     (* Datenbaustein Testen *)
     #rTEST_DB := TEST_DB(DB_NUMBER := #_pt.DBNr // IN: WORD
                        ,DB_LENGTH => #DB_LENGTH // OUT: WORD
                        ,WRITE_PROT => #WRITE_PROT // OUT: BOOL
                        ); // INT
     (* Ende wenn Test-DB <> 0 = Fehler *)
     IF #rTEST_DB <> 0 THEN RETURN; END_IF;
     (* Ende wenn DB zu klein *) 
     IF WORD_TO_INT(#DB_LENGTH)/4 < #size THEN RETURN; END_IF;

     #Adr := DWORD_TO_INT(SHR(IN:=SHL(IN:=#_pt.Adr,N:=8),N:=11));

     (* at first we calualte the arithmetic average of the array *)

     #stop := (#size - 1) / 1;     // (size -SIZEOF(pt)) / SIZEOF(pt);
     #avg := DWORD_TO_REAL(WORD_TO_BLOCK_DB(#_pt.DBNr).DD(#Adr+0));
     FOR #i := 1 TO #stop DO
         #avg := #avg + DWORD_TO_REAL(WORD_TO_BLOCK_DB(#_pt.DBNr).DD(#Adr+#i*4));
     END_FOR;
     #avg := #avg / (#stop + 1);

     (* in a second run we calculate the variance of the array *)

     #_var := (DWORD_TO_REAL(WORD_TO_BLOCK_DB(#_pt.DBNr).DD(#Adr+0)) - #avg) ** 2;
     FOR #i := 1 TO #stop DO
         #_var := #_var + ((DWORD_TO_REAL(WORD_TO_BLOCK_DB(#_pt.DBNr).DD(#Adr+#i*4)) - #avg) ** 2);
     END_FOR;
     #_var := #_var / #stop;

     (* standard deviation is simply the square root of the variance *)

     #sdv := SQRT(#_var);

   (*
   (* standard deviation is simply the square root of the variance *)

   array_sdv := SQRT(array_var(pt, size));
   *)

   (* revision history
   hm  1.4.2007        rev 1.0
       function created

   hm  16. mar. 2008   rev 1.1
       changed type of input size to uint

   *)
END_FUNCTION_BLOCK

FUNCTION_BLOCK "ARRAY_SPR"   // FB18, SCL
TITLE = ARRAY_SPR
{ S7_Optimized_Access := 'FALSE' }
AUTHOR : hugo
FAMILY : ARFUNCT
NAME : AR_SPR
VERSION : 1.1
// this function will calculate the spread of a given array.
// the function needs to be called:    array_spr(adr("array"),sizeof("array"));
// for example: spread of [12,0,4,1,7] is 12 - 0 = 12.
// because this function works with pointers its very time efficient and it needs no extra memory.
   VAR_INPUT
      pt : Pointer;
      _pt AT pt : Struct
         DBNr : Word;
         Adr : DWord;
      END_STRUCT;
      size : Int;
   END_VAR
   VAR_OUTPUT
      spr : Real;
   END_VAR
   VAR_TEMP
      i : Int;
      stop : Int;
      array_max : Real;
      array_min : Real;
      Adr : Int;
      DB_LENGTH : Word;
      WRITE_PROT : Bool;
      rTEST_DB : Int;
   END_VAR
BEGIN


     (* Datenbaustein Testen *)
     #rTEST_DB := TEST_DB(DB_NUMBER := #_pt.DBNr // IN: WORD
                        ,DB_LENGTH => #DB_LENGTH // OUT: WORD
                        ,WRITE_PROT => #WRITE_PROT // OUT: BOOL
                        ); // INT
     (* Ende wenn Test-DB <> 0 = Fehler *)
     IF #rTEST_DB <> 0 THEN RETURN; END_IF;
     (* Ende wenn DB zu klein *) 
     IF WORD_TO_INT(#DB_LENGTH)/4 < #size THEN RETURN; END_IF;

     #Adr := DWORD_TO_INT(SHR(IN:=SHL(IN:=#_pt.Adr,N:=8),N:=11));

     (* Berechnung *)
     #stop := (#size - #size / #size);
     #array_min := DWORD_TO_REAL(WORD_TO_BLOCK_DB(#_pt.DBNr).DD(#Adr+0));
     #array_max := DWORD_TO_REAL(WORD_TO_BLOCK_DB(#_pt.DBNr).DD(#Adr+0));
     FOR #i := 1 TO #stop DO
         IF DWORD_TO_REAL(WORD_TO_BLOCK_DB(#_pt.DBNr).DD(#Adr+#i*4)) > #array_max THEN 
             #array_max := DWORD_TO_REAL(WORD_TO_BLOCK_DB(#_pt.DBNr).DD(#Adr+#i*4));
         ELSIF DWORD_TO_REAL(WORD_TO_BLOCK_DB(#_pt.DBNr).DD(#Adr+#i*4)) < #array_min THEN 
             #array_min := DWORD_TO_REAL(WORD_TO_BLOCK_DB(#_pt.DBNr).DD(#Adr+#i*4));
         END_IF;
     END_FOR;
     #spr := #array_max - #array_min;

   (* revision history
   hm  2. oct. 2006    rev 1.0
       original version

   hm  16. mar. 2008   rev 1.1
       changed type of input size to uint

   *)
END_FUNCTION_BLOCK

FUNCTION_BLOCK "ARRAY_SUM"   // FB19, SCL
TITLE = ARRAY_SUM
{ S7_Optimized_Access := 'FALSE' }
AUTHOR : hugo
FAMILY : ARFUNCT
NAME : AR_SUM
VERSION : 1.1
// this function will calculate the sum of a given array.
   VAR_INPUT
      pt : Pointer;
      _pt AT pt : Struct
         DBNr : Word;
         Adr : DWord;
      END_STRUCT;
      size : Int;
   END_VAR
   VAR_OUTPUT
      sum : Real;
   END_VAR
   VAR_TEMP
      i : Int;
      Adr : Int;
      DB_LENGTH : Word;
      WRITE_PROT : Bool;
      rTEST_DB : Int;
   END_VAR
BEGIN


     (* Datenbaustein Testen *)
     #rTEST_DB := TEST_DB(DB_NUMBER := #_pt.DBNr // IN: WORD
                        ,DB_LENGTH => #DB_LENGTH // OUT: WORD
                        ,WRITE_PROT => #WRITE_PROT // OUT: BOOL
                        ); // INT
     (* Ende wenn Test-DB <> 0 = Fehler *)
     IF #rTEST_DB <> 0 THEN RETURN; END_IF;
     (* Ende wenn DB zu klein *) 
     IF WORD_TO_INT(#DB_LENGTH)/4 < #size THEN RETURN; END_IF;

     #Adr := DWORD_TO_INT(SHR(IN:=SHL(IN:=#_pt.Adr,N:=8),N:=11));

     (* Berechnung *)
     #sum := DWORD_TO_REAL(WORD_TO_BLOCK_DB(#_pt.DBNr).DD(#Adr+0));
     FOR #i := 1 TO #size-1 DO
         #sum := #sum + DWORD_TO_REAL(WORD_TO_BLOCK_DB(#_pt.DBNr).DD(#Adr+#i*4));
     END_FOR;

   (* revision history
   hm  2. oct. 2006    rev 1.0
       function created

   hm  16. mar. 2008   rev 1.1
       changed type of input size to uint

   *)
END_FUNCTION_BLOCK

FUNCTION_BLOCK "ARRAY_TREND"   // FB20, SCL
TITLE = ARRAY_TREND
{ S7_Optimized_Access := 'FALSE' }
AUTHOR : hugo
FAMILY : ARFUNCT
NAME : AR_TREND
VERSION : 1.3
// this function will calculate the trend of a given array.
// trend will calculate the avg of the first half of the array and then the avg of the second half, trend = avg2 - avg1.
// for example:  [0,1,4,5,3,4,6,3] = 4 - 2.5 = 1.5
// the function needs to be called:    array_trend(adr("array"),sizeof("array"));
// because this function works with pointers its very time efficient and it needs no extra memory.
// 
// uses: EVEN [FC76]
   VAR_INPUT
      pt : Pointer;
      _pt AT pt : Struct
         DBNr : Word;
         Adr : DWord;
      END_STRUCT;
      size : Int;
   END_VAR
   VAR_OUTPUT
      trend : Real;
   END_VAR
   VAR_TEMP
      i : Int;
      stop : Int;
      stop2 : Int;
      x : Real;
      Adr : Int;
      DB_LENGTH : Word;
      WRITE_PROT : Bool;
      rTEST_DB : Int;
   END_VAR
BEGIN


   (* Datenbaustein Testen *)
   #rTEST_DB := TEST_DB(DB_NUMBER := #_pt.DBNr, DB_LENGTH => #DB_LENGTH, WRITE_PROT => #WRITE_PROT);
   (* Ende wenn Test-DB <> 0 = Fehler *)
   IF #rTEST_DB <> 0 THEN RETURN; END_IF;
   (* Ende wenn DB zu klein *) 
   IF WORD_TO_INT(#DB_LENGTH)/4 < #size THEN RETURN; END_IF;

   #Adr := DWORD_TO_INT(SHR(IN:=SHL(IN:=#_pt.Adr,N:=8),N:=11));

   #stop := #size - 1;
   #stop2 := #stop / 2;
   FOR #i := 0 TO #stop2 DO #x := #x - DWORD_TO_REAL(WORD_TO_BLOCK_DB(#_pt.DBNr).DD(#Adr+#i*4)); END_FOR;
   IF "EVEN"(#stop) THEN
       FOR #i := #stop2 TO #stop DO #x := #x + DWORD_TO_REAL(WORD_TO_BLOCK_DB(#_pt.DBNr).DD(#Adr+#i*4)); END_FOR;
   ELSE
       FOR #i := #stop2 + 1 TO #stop DO #x := #x + DWORD_TO_REAL(WORD_TO_BLOCK_DB(#_pt.DBNr).DD(#Adr+#i*4)); END_FOR;
   END_IF;
   #trend := #x / INT_TO_REAL(#stop2 + 1);


   (* revision history
   hm  2 oct 2007  rev 1.0
       original version

   hm  12 dec 2007 rev 1.1
       changed code for better performance

   hm  16. mar. 2008   rev 1.2
       changed type of input size to uint

   hm  10. mar. 2009   rev 1.3
       added type conversions for compatibility reasons
   *)
END_FUNCTION_BLOCK

FUNCTION_BLOCK "ARRAY_VAR"   // FB21, SCL
TITLE = ARRAY_VAR
{ S7_Optimized_Access := 'FALSE' }
AUTHOR : hugo
FAMILY : ARFUNCT
NAME : AR_VAR
VERSION : 1.3
// this function will calculate the variance of a given array.
// the function needs to be called:    array_var(adr("array"),sizeof("array"));
// because this function works with pointers its very time efficient and it needs no extra memory.
   VAR_INPUT
      pt : Pointer;
      _pt AT pt : Struct
         DBNr : Word;
         Adr : DWord;
      END_STRUCT;
      size : Int;
   END_VAR
   VAR_OUTPUT
      _var : Real;
   END_VAR
   VAR_TEMP
      i : Int;
      stop : Int;
      avg : Real;
      Adr : Int;
      DB_LENGTH : Word;
      WRITE_PROT : Bool;
      rTEST_DB : Int;
   END_VAR
BEGIN


   (* Datenbaustein Testen *)
   #rTEST_DB := TEST_DB(DB_NUMBER := #_pt.DBNr, DB_LENGTH => #DB_LENGTH, WRITE_PROT => #WRITE_PROT);
   (* Ende wenn Test-DB <> 0 = Fehler *)
   IF #rTEST_DB <> 0 THEN RETURN; END_IF;
   (* Ende wenn DB zu klein *) 
   IF WORD_TO_INT(#DB_LENGTH)/4 < #size THEN RETURN; END_IF;

   #Adr := DWORD_TO_INT(SHR(IN:=SHL(IN:=#_pt.Adr,N:=8),N:=11));

   (* at first we calualte the arithmetic average of the array *)

   #stop := #size - 1;
   #avg := DWORD_TO_REAL(WORD_TO_BLOCK_DB(#_pt.DBNr).DD(#Adr+0));
   FOR #i := 1 TO #stop DO
       #avg := #avg + DWORD_TO_REAL(WORD_TO_BLOCK_DB(#_pt.DBNr).DD(#Adr+#i*4));
   END_FOR;
   #avg := #avg / (#stop + 1);

   (* in a second run we calculate the variance of the array *)

   #_var := (DWORD_TO_REAL(WORD_TO_BLOCK_DB(#_pt.DBNr).DD(#Adr+0)) - #avg) * (DWORD_TO_REAL(WORD_TO_BLOCK_DB(#_pt.DBNr).DD(#Adr+0)) - #avg);
   FOR #i := 1 TO #stop DO
       #_var := #_var + (DWORD_TO_REAL(WORD_TO_BLOCK_DB(#_pt.DBNr).DD(#Adr+#i*4)) - #avg) * (DWORD_TO_REAL(WORD_TO_BLOCK_DB(#_pt.DBNr).DD(#Adr+#i*4)) - #avg);
   END_FOR;
   #_var := #_var / INT_TO_REAL(#stop);


   (* revision history
   hm  1.4.2007    rev 1.0
       function created

   hm  12.12.2007  rev 1.1
       changed code for better performance

   hm  16. mar. 2008   rev 1.2
       changed type of input size to uint

   hm  10. mar. 2009   rev 1.3
       added type conversions for compatibility reasons
   *)
END_FUNCTION_BLOCK

FUNCTION_BLOCK "IS_SORTED"   // FB22, SCL
TITLE = IS_SORTED
{ S7_Optimized_Access := 'FALSE' }
AUTHOR : hugo
FAMILY : ARFUNCT
NAME : ARSORTED
VERSION : 1.1
// this function will return true if the given array is sorted in an ascending order.
// the function needs to be called:    array_sorted(adr("array"),sizeof("array"));
// because this function works with pointers its very time efficient and it needs no extra memory.
   VAR_INPUT
      pt : Pointer;
      _pt AT pt : Struct
         DBNr : Word;
         Adr : DWord;
      END_STRUCT;
      size : Int;
   END_VAR
   VAR_OUTPUT
      SORTED : Bool;
   END_VAR
   VAR
      stop : Int;
      i : Int;
      Adr : Int;
      DB_LENGTH : Word;
      WRITE_PROT : Bool;
      rTEST_DB : Int;
   END_VAR
BEGIN


   #SORTED := FALSE;

   (* Datenbaustein Testen *)
   #rTEST_DB := TEST_DB(DB_NUMBER := #_pt.DBNr // IN: WORD
                      ,DB_LENGTH => #DB_LENGTH // OUT: WORD
                      ,WRITE_PROT => #WRITE_PROT // OUT: BOOL
                      ); // INT
   (* Ende wenn Test-DB <> 0 = Fehler *)
   IF #rTEST_DB <> 0 THEN RETURN; END_IF;
   (* Ende wenn DB zu klein *) 
   IF WORD_TO_INT(#DB_LENGTH)/4 < #size THEN RETURN; END_IF;

   #Adr := DWORD_TO_INT(SHR(IN:=SHL(IN:=#_pt.Adr,N:=8),N:=11));

   #stop := #size - 2;   //WORD_TO_INT(SHR(IN:=INT_TO_WORD(size),N:=2))-2;
   FOR #i := 0 TO #stop DO
       IF DWORD_TO_REAL(WORD_TO_BLOCK_DB(#_pt.DBNr).DD(#Adr+#i*4)) > DWORD_TO_REAL(WORD_TO_BLOCK_DB(#_pt.DBNr).DD(#Adr+(#i+1)*4)) THEN
           #SORTED := FALSE;
           RETURN;
       END_IF;
   END_FOR;
   #SORTED := TRUE;

   (* revision history

   hm  29. mar. 2008   rev 1.0
       original version

   hm  4. apr. 2008    rev 1.1
       added type conversion to avoid warnings under codesys 3.0
   *)
END_FUNCTION_BLOCK

FUNCTION_BLOCK "STIME"   // FB64, SCL
TITLE = STIME
{ S7_Optimized_Access := 'FALSE' }
AUTHOR : dalbi
FAMILY : MEASURE
NAME : STIME
VERSION : 1.4
// this function block makes sure that the timer of a siemens sps counts from 0 - 2^32-1.
   VAR_OUTPUT
      tx : DWord;
      at_tx AT tx : Array[0..31] of Bool;
   END_VAR
   VAR
      last_time : DWord;
      bit31 : Bool;
      init : Bool := TRUE;
   END_VAR
   VAR_TEMP
      TOP_SI : Struct
         EV_CLASS : Byte;
         EV_NUM : Byte;
         PRIORITY : Byte;
         NUM : Byte;
         TYP2_3 : Byte;
         TYP1 : Byte;
         ZI1 : Word;
         ZI2_3 : DWord;
      END_STRUCT;
      START_UP_SI : Struct
         EV_CLASS : Byte;
         EV_NUM : Byte;
         PRIORITY : Byte;
         NUM : Byte;
         TYP2_3 : Byte;
         TYP1 : Byte;
         ZI1 : Word;
         ZI2_3 : DWord;
      END_STRUCT;
      ERR : Int;
   END_VAR
BEGIN


   (* this FB is only necessary for siemens sps
   the siemens sps timer counts from 0 to 2^31-1 and starts at 0 sfter overrun.
   this means that the bit 31 (the highest bit ) will never be used and therefore
   a problem arises when t2 - t1 is checked.
   t2 - t1 is always valid also in an timer overrun situation where the time t1 is very high and t2 is very low.
   the result of the subtraction t2 - t1 however is still valid.
   this calculation does not work for soiemens because the highest bit is not used.

   this module stores the highest bit, changes the highest bit at every overrun occurence and stuffs ther highest bit in the output.
   the output is then used by t_plc_us and t_plc_ms.

   the correction needs and fb and not a function because the value of the highest bit has to be stored.

   do never use this function block in a codesys environment. the timer in codesys is correct and runs from 0 to 2^32-1
   *)

   (* read actual startup info *)
   (* OB1_SCAN_1  BYTE  -  B#16#01: Abschluss des Neustarts (Warmstarts)
                        -  B#16#02: Abschluss des Wiederanlaufs
                        -  B#16#03: Abschluss des freien Zyklus
                        -  B#16#04: Abschluss des Kaltstarts
                        -  B#16#05: Erster OB 1-Zyklus der neuen Master-CPU nach 
                                    Master-Reserve-Umschaltung und STOP des 
                                    bisherigen Masters *)

   #ERR := RD_SINFO (TOP_SI => #TOP_SI, START_UP_SI => #START_UP_SI);

   (* reset last_time on system startup *)
   IF #TOP_SI.EV_NUM = 1 OR #TOP_SI.EV_NUM = 2 OR #TOP_SI.EV_NUM = 4 OR NOT #init THEN 
       #last_time := 0;
       #bit31 := false;
       #init := true;
   END_IF;

   (* read the system timer *)
   #tx := DINT_TO_DWORD(T_CONV(TIME_TCK()));

   (* check for overrun *)
   IF DWORD_TO_DINT(#tx) < DWORD_TO_DINT(#last_time) THEN
       (* an overrun has occured, change the value of the highest bit *)
       #bit31 := NOT #bit31;
   END_IF;

   (* stuff the highest bit into the timer value *)
   #at_tx[7] := #bit31;

   (* remember the last system time for the next overrun check *)
   #last_time := #tx;


   (* revision history
   DA  14.9.2007 rev 1.0
     original version

   DA  24.2.2008 rev 1.1
     added self reset on system startup

   DA   2.5.2008 rev 1.2
     corect a problem running under OB35

   DA  12.3.2009 rev 1.3
     corect a problem run on different CPUs

   DA  22.12.2009 rev 1.4
     corect a problem on startup
   *)
END_FUNCTION_BLOCK

FUNCTION "T_PLC_MS" : DWord   // FC64, SCL
TITLE = T_PLC_MS
{ S7_Optimized_Access := 'FALSE' }
AUTHOR : hugo
FAMILY : MEASURE
NAME : T_PLC_MS
VERSION : 1.2
// T_PLC_MS reads the internal PLC timer and return the time, it has the advantage to be able to set a debug mode 
// and speed up the counter to test the plc timer overrun which occurs every 50 days respectively 25 days at siemens S7
// this routine also allows to correct the behavior of s7 where the internal plc counter will not count all 32 bits.
// 
// uses: STIME [FB64],IDB_STIME [DB64]
BEGIN


   "IDB_STIME"(); 
   #T_PLC_MS := "IDB_STIME".tx; 
   (* hier muss die korrektur für step7 stattfinden
   plctime muss den vollen wertebereich von time ausnutzen:
   wenn bei step7 time -24tage bis plus 24 tage ist dann muss der timer auch beim überlauf auf -24tage springen 
   und auf keinen fall auf 0 !!!!
   für siemens muss ein weiterer fb im main eingebunden werden der sicherstellt das alle 32 bits durchgezählt werden.
   es kann nur ein fb sein den er muss sich das oberste (32te) bit merken.
   oder etwa spring s7 bei überlauf auf -24 tage????? dann wäre keine korrektur nötig.
   *)
   IF "debug" THEN
       #T_PLC_MS := DINT_TO_DWORD((DWORD_TO_DINT(SHL(IN:=#T_PLC_MS,N:="N") OR SHL(IN:=DWORD#1,N:="N"))-1) + DWORD_TO_DINT("offset_1"));
   END_IF;


   (* revision history
   hm  14.9.2007   rev 1.0
       original version

   hm  12. nov 2007    rev 1.1
       added temporaray variable tx because some compilers could not handle time() as an argument

   hm  16. nov. 2008   rev 1.2
       initialized constants with 0 for compatibility reasons
   *)
END_FUNCTION

FUNCTION "EVEN" : Bool   // FC76, SCL
TITLE = EVEN
{ S7_Optimized_Access := 'FALSE' }
AUTHOR : hugo
FAMILY : MATH
NAME : EVEN
VERSION : 1.2
// this function chacks an input for even value
// the output is true if the input is even.
   VAR_INPUT
      in : DInt;
   END_VAR
   VAR_TEMP
      tIN : DInt;
      _IN AT tIN : Array[0..31] of Bool;
   END_VAR
BEGIN


   #tIN := #in;
   #EVEN := NOT #_IN[24]; //EVEN := NOT in.0;

   (* revision history
   hm  1. oct 2006 rev 1.0
     ORIGINAL VERSION

   hm  01.12.2007  rev 1.1
     changed code for improved performance

   hm  21. mar. 2008 rev 1.2
     changed type of input IN from INT to DINT
   *)
END_FUNCTION

FUNCTION "FRACT" : Real   // FC83, SCL
TITLE = FRACT
{ S7_Optimized_Access := 'FALSE' }
AUTHOR : hugo
FAMILY : MATH
NAME : FRACT
VERSION : 1.3
// this function returns the fraction of a real number
// fract(3.14) = 0.14
   VAR_INPUT
      x : Real;
   END_VAR
BEGIN


   IF ABS(#x) < 2.0E9 THEN
       #FRACT := #x - DINT_TO_REAL(TRUNC(#x));
   ELSE
       #FRACT := 0.0;
   END_IF;


   (* revision history
   hm  4. aug 2006 rev 1.0
       original version

   hm  11. mar 2008    rev 1.1
       added dint_to_real for compatibility reasons
       now returns 0 for number > 2e9
       changed input to x

   hm  21. mar. 2008   rev 1.2
       use D_trunc instead of TRUNC for compatibility reasons

   hm  10. mar. 2009   rev 1.3
       real constants updated to new systax using dot

   *)
END_FUNCTION

FUNCTION "RDM" : Real   // FC101, SCL
TITLE = RDM
{ S7_Optimized_Access := 'FALSE' }
AUTHOR : hugo
FAMILY : MATH
NAME : RDM
VERSION : 1.9
// this function calculates a pseudo random number
// to generate the number it reads the sps timer and calculates a random number between 0 and 1:
// in order to use rdm more then once within one sps cycle it need to be called with different seed numbers LAST.
//  
// uses: T_PLC_MS [FC64]
//       STIME [FB64],IDB_STIME [DB64]
//       BIT_COUNT [FC291]
//       FRACT [FC83]
   VAR_INPUT
      last : Real;
   END_VAR
   VAR_TEMP
      tn : DWord;
      _tn AT tn : Array[0..31] of Bool;
      tc : Int;
   END_VAR
BEGIN


   #tn := "T_PLC_MS"();
   #tc := "BIT_COUNT"(#tn);
   #_tn[7] := #_tn[26];  //tn.31 := tn.2;
   #_tn[6] := #_tn[29];  //tn.30 := tn.5;
   #_tn[5] := #_tn[28];  //tn.29 := tn.4;
   #_tn[4] := #_tn[25];  //tn.28 := tn.1;
   #_tn[3] := #_tn[24];  //tn.27 := tn.0;
   #_tn[2] := #_tn[31];  //tn.26 := tn.7;
   #_tn[1] := #_tn[30];  //tn.25 := tn.6;
   #_tn[0] := #_tn[27];  //tn.24 := tn.3;
   #tn := ROL(IN:=#tn,N:="BIT_COUNT"(#tn)) AND 16#7FFFFFFF OR 16#40000001;  // OR 16#80000001
   #tn := DINT_TO_DWORD(DWORD_TO_DINT(#tn) MOD 71474513 + #tc + 77);
   #RDM := "FRACT"(DINT_TO_REAL(DWORD_TO_DINT(#tn)) / 10000000.0 * ("E"- LIMIT(MN:=0.0,IN:=#last,MX:=1.0)));


   (*
   pt := ADR(temp);
   pt^ := (T_PLC_MS() AND 16#007FFFFF) OR 16#3D000000;
   RDM := fract(modR(temp*e+pi1, PI1-last) + modR(temp*PI1+e + last,e-last));
   *)

   (* revision history
   hm      16. jan 2007        rev 1.0
       original version

   hm      11. nov 2007        rev 1.1
       changed time() into t_plc_ms()

   hm      20. nov 2007        rev 1.2
       changed code of temp calculation to avoid overflow in modr due to resuclt would not fit DINT for high timeer values

   hm      5. jan 2008     rev 1.3
       changed calculation of temp to avoid problem with high values of t_plc_ms

   hm      2. feb 2008     rev 1.4
       changed algorithm to avoind non iec functions and guarantee more randomness

   hm  10. mar. 2008       rev 1.5
       make sure last will be between 0 and 1 to avoid invalid results

   hm  16. mar. 2008       rev 1.6
       added conversion for tc to avoid warnings under codesys 3.0

   hm  18. may. 2008       rev 1.7
       changed constant E to E1

   hm  18. oct. 2008       rev 1.8
       using math constants

   hm  10. mar. 2009       rev 1.9
       real constants updated to new systax using dot

   *)
END_FUNCTION

FUNCTION "RDM2" : Int   // FC102, SCL
TITLE = RDM2
{ S7_Optimized_Access := 'FALSE' }
AUTHOR : hugo
FAMILY : MATH
NAME : RDM2
VERSION : 1.1
// this function calculates an integer pseudo random number
// the random number will be in the range of low <= rdm2 <= high.
// 
// uses: RDM [FC101]
//       T_PLC_MS [FC64] 
//       STIME [FB64],IDB_STIME [DB64] 
//       BIT_COUNT [FC291] 
//       FRACT [FC83]
   VAR_INPUT
      last : Int;
      low : Int;
      high : Int;
   END_VAR
BEGIN


   #RDM2 := REAL_TO_INT(DINT_TO_REAL(TRUNC("RDM"("FRACT"(#last*"PI")) * (#high - #low + 1)) + #low));

   (* revision history
   hm      29. feb 2008        rev 1.0
       original version

   hm      18. oct. 2008       rev 1.1
       using math constants

   *)
END_FUNCTION

FUNCTION "SQRTN" : Real   // FC112, SCL
TITLE = SQRTN
{ S7_Optimized_Access := 'FALSE' }
AUTHOR : hugo
FAMILY : MATH
NAME : SQRTN
VERSION : 1.3
// this function calculates the nth root function of X according to the formula sqrtn = x^(1/n).
   VAR_INPUT
      X : Real;
      N : Int;
   END_VAR
BEGIN


   IF #N > 0 THEN
       #SQRTN := EXP(LN(#X) / INT_TO_REAL(#N));
   ELSE
       #SQRTN := 0.0;
   END_IF;


   (* revision history
   hm      12 jan 2007 rev 1.0
       original version

   hm      2. dec 2007 rev 1.1
       changed code for better performance

   hm      11. mar 2008    rev 1.2
       added result 0 for compatibility reasons

   hm 10. mar. 2009    rev 1.3
       added type conversions for compatibility reasons

   *)
END_FUNCTION

FUNCTION "BIT_COUNT" : Int   // FC291, SCL
TITLE = BIT_COUNT
{ S7_Optimized_Access := 'FALSE' }
AUTHOR : hugo
FAMILY : GATE
NAME : BITCT
VERSION : 1.1
// BIT_COUNT counts the amount True of bits in a dword.
// for exabple: bit_count(3) returns 2 because two bits (bits 0 and 1) are true and all others are false.
   VAR_INPUT
      IN : DWord;
   END_VAR
   VAR_TEMP
      temp : DWord;
      attemp AT temp : Array[0..31] of Bool;
   END_VAR
BEGIN


     #BIT_COUNT := 0;
     #temp := #IN;

     WHILE DWORD_TO_DINT(#temp) <> 0 DO
       IF #attemp[24] THEN #BIT_COUNT := #BIT_COUNT +1; END_IF;
       #temp := SHR(IN:=#temp,N:=1);
     END_WHILE;

   (* revision history
   5.7.2007  rev 1.0    original version

   10.9.2007  rev 1.1    hm
     changed algorithm for better performace
     the execution time has reduced by a factor of 5
     deleted unused variable temp
   *)
END_FUNCTION

// ===== PLC "Mathematical Complex"  Unspecific CPU S7 300 =====

VAR_GLOBAL CONSTANT   // PLC tag table "STEP7 classic symbols"
   "PI1" : Real := 3.14159265358979323846264338327950288;
   "PI05" : Real := 1.5707963267949;
END_VAR

TYPE "COMPLEX"
VERSION : 0.0
   STRUCT
      re : Real;
      im : Real;
   END_STRUCT;
END_TYPE

FUNCTION "ATAN2" : Real   // FC58, SCL
TITLE = ATAN2
{ S7_Optimized_Access := 'FALSE' }
AUTHOR : hugo
FAMILY : MATH
NAME : ATAN2
VERSION : 1.2
// this function calculates the angle in a coordinate system in rad.
   VAR_INPUT
      Y : Real;
      X : Real;
   END_VAR
BEGIN


   IF #X > 0.0 THEN
       #ATAN2 := ATAN(#Y/#X);
   ELSIF #X < 0.0 THEN
       IF #Y >= 0.0 THEN
           #ATAN2 := ATAN(#Y/#X) + "PI1";
       ELSE
           #ATAN2 := ATAN(#Y/#X) - "PI1";
       END_IF;
   ELSIF #Y > 0.0 THEN
       #ATAN2 := "PI05";
   ELSIF #Y < 0.0 THEN
       #ATAN2 := -"PI05";
   ELSE
       #ATAN2 := 0.0;
   END_IF;


   (* revision history
   hm  20.  apr. 2008  rev 1.0
       original version

   hm  18. oct. 2008   rev 1.1
       changed to use math constants

   hm  10. mar. 2009   rev 1.2
       real constants updated to new systax using dot

   *)
END_FUNCTION

FUNCTION "COSH" : Real   // FC69, SCL
TITLE = COSH
{ S7_Optimized_Access := 'FALSE' }
AUTHOR : hugo
FAMILY : MATH
NAME : COSH
VERSION : 1.3
// this function calculates the cos hyperbolicus
   VAR_INPUT
      X : Real;
   END_VAR
   VAR_TEMP
      t : Real;
   END_VAR
BEGIN


   #t := EXP(#X);
   #COSH := (1.0 / #t + #t) * 0.5;


   (* revision histroy
   hm  12.1.2007   rev 1.0
       original version

   hm  1.12.2007   rev 1.1
       changed code to improve performance

   hm  5. jan 2008   rev 1.2
       further performance improvement

   hm  10. mar. 2009   rev 1.3
       real constants updated to new systax using dot
   *)
END_FUNCTION

FUNCTION "HYPOT" : Real   // FC89, SCL
TITLE = HYPOT
{ S7_Optimized_Access := 'FALSE' }
AUTHOR : hugo
FAMILY : MATH
NAME : HYPOT
VERSION : 1.0
// this function calculates the pythagorean function
   VAR_INPUT
      X : Real;
      Y : Real;
   END_VAR
BEGIN


     #HYPOT := SQRT(#X*#X + #Y*#Y);


   (* revision history
   hm  21. feb 2008  rev 1.0
     original version

   *)
END_FUNCTION

FUNCTION "SGN" : Int   // FC106, SCL
TITLE = SGN
{ S7_Optimized_Access := 'FALSE' }
AUTHOR : hugo
FAMILY : MATH
NAME : SGN
VERSION : 1.1
// sgn returns 0 when X = 0 , -1 when X < 1 and +1 when X > 1
   VAR_INPUT
      X : Real;
   END_VAR
BEGIN


     IF #X > 0.0 THEN
       #SGN := 1;
     ELSIF #X < 0.0 THEN
       #SGN := -1;
     ELSE
       #SGN := 0;
     END_IF;

   (* revision histroy
   hm  16. oct 2007  rev 1.0
     original version

   hm  11. nov 2007  rev 1.1
     changed type of function from real to int
   *)
END_FUNCTION

FUNCTION "SINH" : Real   // FC111, SCL
TITLE = SINH
{ S7_Optimized_Access := 'FALSE' }
AUTHOR : hugo
FAMILY : MATH
NAME : SINH
VERSION : 1.3
// this function calculates the sin hyperbolicus
   VAR_INPUT
      X : Real;
   END_VAR
BEGIN


   IF ABS(#X) < 2.0E-3 THEN
       #SINH := #X;
   ELSE
       #SINH := (EXP(#X) - EXP(-#X)) * 0.5;
   END_IF;

   (* revision history
   hm  12.1.2007   rev 1.0
       original version

   hm  1.12.2007   rev 1.1
       changed code to improve performance

   hm  5. jan 2008 rev 1.2
       further performance improvement

   hm  11. mar 2008    rev 1.3
       improved accuracy around 0

   *)
END_FUNCTION

FUNCTION "CABS" : Real   // FC117, SCL
TITLE = CABS
{ S7_Optimized_Access := 'FALSE' }
AUTHOR : hugo
FAMILY : CMATH
NAME : CABS
VERSION : 1.0
// this function the aboslute value of a complex number
//  
// uses: COMPLEX [UDT2]
//       HYPOT [FC89]
   VAR_INPUT
      X : "COMPLEX";
   END_VAR
BEGIN


     #CABS := "HYPOT"(X:=#X.re,Y:=#X.im);


   (* revision history
   hm  21. feb 2008  rev 1.0
     original version

   *)
END_FUNCTION

FUNCTION "CACOS" : "COMPLEX"   // FC118, SCL
TITLE = CACOS
{ S7_Optimized_Access := 'FALSE' }
AUTHOR : hugo
FAMILY : CMATH
NAME : CACOS
VERSION : 1.0
// this function calculates the arcus cosinus function of a complex number
// 
// uses: COMPLEX [UDT2]
//       CACOSH [FC119]
//       CSQRT [FC139] 
//       HYPOT [FC89]
//       SGN [FC106]
//       CLOG [FC132] 
//       ATAN2 [FC58]
   VAR_INPUT
      X : "COMPLEX";
   END_VAR
   VAR_TEMP
      Y : "COMPLEX";
      temp_X : "COMPLEX";
      temp_complex : "COMPLEX";
   END_VAR
BEGIN


     #temp_X := #X;

     #Y := "CACOSH"(#temp_X);
     #temp_complex.re := #Y.im;
     #temp_complex.im := -#Y.re;

     #CACOS := #temp_complex;


   (* revision history
   hm  21. feb 2008  rev 1.0
     original version


   *)
END_FUNCTION

FUNCTION "CACOSH" : "COMPLEX"   // FC119, SCL
TITLE = CACOSH
{ S7_Optimized_Access := 'FALSE' }
AUTHOR : hugo
FAMILY : CMATH
NAME : CACOSH
VERSION : 1.0
// this function calculates the hyperbolic arcus cosinus function of a complex number
// 
// uses: COMPLEX [UDT2]
//       CSQRT [FC139]
//       HYPOT [FC89] 
//       SGN [FC106] 
//       CLOG [FC132]
//       ATAN2 [FC58]
   VAR_INPUT
      X : "COMPLEX";
   END_VAR
   VAR_TEMP
      Y : "COMPLEX";
      temp_complex : "COMPLEX";
   END_VAR
BEGIN


     #Y.re := (#X.re - #X.im)*(#X.re + #X.im) - 1.0;
     #Y.im := 2.0 * #X.re * #X.im;
     #Y    := "CSQRT"(#Y);
     #Y.re := #Y.re + #X.re;
     #Y.im := #Y.im + #X.im;
     #temp_complex := "CLOG"(#Y);

     #CACOSH := #temp_complex;


   (* revision history
   hm  21. feb 2008  rev 1.0
     original version


   *)
END_FUNCTION

FUNCTION "CADD" : "COMPLEX"   // FC120, SCL
TITLE = CADD
{ S7_Optimized_Access := 'FALSE' }
AUTHOR : hugo
FAMILY : CMATH
NAME : CADD
VERSION : 1.0
// this function add two complex numbers
// 
// uses: COMPLEX [UDT2]
   VAR_INPUT
      X : "COMPLEX";
      Y : "COMPLEX";
   END_VAR
   VAR_TEMP
      temp_CADD : "COMPLEX";
   END_VAR
BEGIN


     #temp_CADD.re := #X.re + #Y.re;
     #temp_CADD.im := #X.im + #Y.im;

     #CADD := #temp_CADD;

   (* revision history
   hm  21. feb 2008  rev 1.0
     original version

   *)
END_FUNCTION

FUNCTION "CARG" : Real   // FC121, SCL
TITLE = CARG
{ S7_Optimized_Access := 'FALSE' }
AUTHOR : hugo
FAMILY : CMATH
NAME : CARG
VERSION : 1.1
// this function calculates the phase angle (argument) of a complex number
// 
// uses: COMPLEX [UDT2]
//       ATAN2 [FC58]
   VAR_INPUT
      X : "COMPLEX";
   END_VAR
BEGIN


     #CARG := "ATAN2"(Y:=#X.im,X:=#X.re);


   (* revision history
   hm  21. feb. 2008   rev 1.0
       original version

   hm  20. apr. 2008   rev 1.1
       use ATAN2 instead of ATAN
   *)
END_FUNCTION

FUNCTION "CASIN" : "COMPLEX"   // FC122, SCL
TITLE = CASIN
{ S7_Optimized_Access := 'FALSE' }
AUTHOR : hugo
FAMILY : CMATH
NAME : CASIN
VERSION : 1.0
// this function calculates the arcus sinus function of a complex number
// 
// uses: COMPLEX [UDT2]
//       CASINH [FC123]
//       CSQRT [FC139] 
//       HYPOT [FC89]
//       SGN [FC106]
//       CLOG [FC132] 
//       ATAN2 [FC58]
   VAR_INPUT
      X : "COMPLEX";
   END_VAR
   VAR_TEMP
      Y : "COMPLEX";
      temp_CASIN : "COMPLEX";
   END_VAR
BEGIN


     #Y.re := -#X.im;
     #Y.im := #X.re;
     #Y := "CASINH"(#Y);
     #temp_CASIN.re := #Y.im;
     #temp_CASIN.im := -#Y.re;

     #CASIN := #temp_CASIN;


   (* revision history
   hm  21. feb 2008  rev 1.0
     original version


   *)
END_FUNCTION

FUNCTION "CASINH" : "COMPLEX"   // FC123, SCL
TITLE = CASINH
{ S7_Optimized_Access := 'FALSE' }
AUTHOR : hugo
FAMILY : CMATH
NAME : CASINH
VERSION : 1.0
// this function calculates the hyperbolic arcus sinus function of a complex number
// 
// uses: COMPLEX [UDT2]
//       CSQRT [FC139]
//       HYPOT [FC89] 
//       SGN [FC106] 
//       CLOG [FC132]
//       ATAN2 [FC58]
   VAR_INPUT
      X : "COMPLEX";
   END_VAR
   VAR_TEMP
      Y : "COMPLEX";
      temp_CASINH : "COMPLEX";
   END_VAR
BEGIN


     #Y.re := (#X.re - #X.im)*(#X.re + #X.im) + 1.0;
     #Y.im := 2.0 * #X.re * #X.im;
     #Y    := "CSQRT"(#Y);
     #Y.re := #Y.re + #X.re;
     #Y.im := #Y.im + #X.im;
     #temp_CASINH  := "CLOG"(#Y);

     #CASINH := #temp_CASINH;


   (* revision history
   hm  21. feb 2008  rev 1.0
     original version


   *)
END_FUNCTION

FUNCTION "CATAN" : "COMPLEX"   // FC124, SCL
TITLE = CATAN
{ S7_Optimized_Access := 'FALSE' }
AUTHOR : hugo
FAMILY : CMATH
NAME : CATAN
VERSION : 1.0
// this function calculates the complex arcus tangens
//  
// uses: COMPLEX [UDT2]
   VAR_INPUT
      X : "COMPLEX";
   END_VAR
   VAR_TEMP
      r2 : Real;
      num : Real;
      den : Real;
      temp_CATAN : "COMPLEX";
   END_VAR
BEGIN


     #r2 := #X.re * #X.re;
     #den := 1.0 - #r2 - #X.im * #X.im;
     #temp_CATAN.re := 0.5 * ATAN(2.0 * #X.re / #den);
     #num := #X.im + 1.0;
     #num := #r2 + #num * #num;
     #den := #X.im - 1.0;
     #den := #r2 + #den * #den;
     #temp_CATAN.im := 0.25 * (LN(#num)-LN(#den));

     #CATAN := #temp_CATAN;

   (* revision history
   hm  21. feb 2008  rev 1.0
     original version


   *)
END_FUNCTION

FUNCTION "CATANH" : "COMPLEX"   // FC125, SCL
TITLE = CATANH
{ S7_Optimized_Access := 'FALSE' }
AUTHOR : hugo
FAMILY : CMATH
NAME : CATANH
VERSION : 1.0
// this function calculates the complex arcus hyperbolic tangens
//  
// uses: COMPLEX [UDT2]
   VAR_INPUT
      X : "COMPLEX";
   END_VAR
   VAR_TEMP
      i2 : Real;
      num : Real;
      den : Real;
      temp_CATANH : "COMPLEX";
   END_VAR
BEGIN


     #i2 := #X.im * #X.im;
     #num := 1.0 + #X.re;
     #num := #i2 + #num * #num;
     #den := 1.0 - #X.re;
     #den := #i2 + #den * #den;
     #temp_CATANH.re := 0.25 * (LN(#num) - LN(#den));
     #den := 1 - #X.re * #X.re - #i2;
     #temp_CATANH.im := 0.5 * ATAN(2.0 * #X.im / #den);

     #CATANH := #temp_CATANH;

   (* revision history
   hm  21. feb 2008  rev 1.0
     original version


   *)
END_FUNCTION

FUNCTION "CCON" : "COMPLEX"   // FC126, SCL
TITLE = CCON
{ S7_Optimized_Access := 'FALSE' }
AUTHOR : hugo
FAMILY : CMATH
NAME : CCON
VERSION : 1.0
// this function calcucates the conjugation of a complex number
// 
// uses: COMPLEX [UDT2]
   VAR_INPUT
      X : "COMPLEX";
   END_VAR
   VAR_TEMP
      temp_CCON : "COMPLEX";
   END_VAR
BEGIN


     #CCON.re := #X.re;
     #CCON.im := -#X.im;

     #CCON := #temp_CCON;

   (* revision history
   hm  21. feb 2008  rev 1.0
     original version

   *)
END_FUNCTION

FUNCTION "CCOS" : "COMPLEX"   // FC127, SCL
TITLE = CCOS
{ S7_Optimized_Access := 'FALSE' }
AUTHOR : hugo
FAMILY : CMATH
NAME : CCOS
VERSION : 1.0
// this function calculates the cosinus function of a complex number
// 
// uses: COMPLEX [UDT2]
//       CCOSH [FC128]
//       COSH [FC69] 
//       SINH [FC111] 
//       CSET [FC136]
   VAR_INPUT
      X : "COMPLEX";
   END_VAR
   VAR_TEMP
      temp_CCOS : "COMPLEX";
   END_VAR
BEGIN


     #temp_CCOS := "CCOSH"("CSET"(RE:=-#X.im,IM:=#X.re));

     #CCOS := #temp_CCOS;

   (* revision history
   hm  21. feb 2008  rev 1.0
     original version

   *)
END_FUNCTION

FUNCTION "CCOSH" : "COMPLEX"   // FC128, SCL
TITLE = CCOSH
{ S7_Optimized_Access := 'FALSE' }
AUTHOR : hugo
FAMILY : CMATH
NAME : CCOSH
VERSION : 1.0
// this function calculates the arcus tangens function of a complex number
// 
// uses: COMPLEX [UDT2]
//       COSH [FC69]
//       SINH [FC111]
   VAR_INPUT
      X : "COMPLEX";
   END_VAR
   VAR_TEMP
      temp_CCOSH : "COMPLEX";
   END_VAR
BEGIN


     #temp_CCOSH.re := "COSH"(#X.re) * COS(#X.im);
     #temp_CCOSH.im := "SINH"(#X.re) * SIN(#X.im);

     #CCOSH := #temp_CCOSH;

   (* revision history
   hm  21. feb 2008  rev 1.0
     original version

   *)
END_FUNCTION

FUNCTION "CDIV" : "COMPLEX"   // FC129, SCL
TITLE = CDIV
{ S7_Optimized_Access := 'FALSE' }
AUTHOR : hugo
FAMILY : CMATH
NAME : CDIV
VERSION : 1.0
// this function divides two complex numbers
// 
// uses: COMPLEX [UDT2]
   VAR_INPUT
      X : "COMPLEX";
      Y : "COMPLEX";
   END_VAR
   VAR_TEMP
      Temp : Real;
      temp_CDIV : "COMPLEX";
   END_VAR
BEGIN


     #Temp := #Y.re * #Y.re + #Y.im * #Y.im;
     #temp_CDIV.re := (#X.re * #Y.re + #X.im * #Y.im) / #Temp;
     #temp_CDIV.im := (#X.im * #Y.re - #X.re * #Y.im) / #Temp;

     #CDIV := #temp_CDIV;

   (* revision history
   hm  21. feb 2008  rev 1.0
     original version

   *)
END_FUNCTION

FUNCTION "CEXP" : "COMPLEX"   // FC130, SCL
TITLE = CEXP
{ S7_Optimized_Access := 'FALSE' }
AUTHOR : hugo
FAMILY : CMATH
NAME : CEXP
VERSION : 1.0
// this function calculates the complex exponent
// 
// uses: COMPLEX [UDT2]
   VAR_INPUT
      X : "COMPLEX";
   END_VAR
   VAR_TEMP
      Temp : Real;
      temp_CEXP : "COMPLEX";
   END_VAR
BEGIN


     #Temp := EXP(#X.re);
     #temp_CEXP.re := #Temp * COS(#X.im);
     #temp_CEXP.im := #Temp * SIN(#X.im);

     #CEXP := #temp_CEXP;

   (* revision history
   hm  21. feb 2008  rev 1.0
     original version

   *)
END_FUNCTION

FUNCTION "CINV" : "COMPLEX"   // FC131, SCL
TITLE = CINV
{ S7_Optimized_Access := 'FALSE' }
AUTHOR : hugo
FAMILY : CMATH
NAME : CINV
VERSION : 1.0
// this function calculates the inverse of a complex numbers (1 / X)
// 
// uses: COMPLEX [UDT2]
   VAR_INPUT
      X : "COMPLEX";
   END_VAR
   VAR_TEMP
      temp : Real;
      temp_CINV : "COMPLEX";
   END_VAR
BEGIN


     #temp := #X.re * #X.re + #X.im * #X.im;
     #temp_CINV.re := #X.re / #temp;
     #temp_CINV.im := -#X.im / #temp;

     #CINV := #temp_CINV;

   (* revision history
   hm  21. feb 2008  rev 1.0
     original version

   *)
END_FUNCTION

FUNCTION "CLOG" : "COMPLEX"   // FC132, SCL
TITLE = CLOG
{ S7_Optimized_Access := 'FALSE' }
AUTHOR : hugo
FAMILY : CMATH
NAME : CLOG
VERSION : 1.0
// this function calculates the complex natural (base e) logarithm
// 
// uses: COMPLEX [UDT2]
//       HYPOT [FC89]
//       ATAN2 [FC58]
   VAR_INPUT
      X : "COMPLEX";
   END_VAR
   VAR_TEMP
      temp_complex : "COMPLEX";
   END_VAR
BEGIN


   #temp_complex.re := LN("HYPOT"(X:=#X.re,Y:=#X.im));
   #temp_complex.im := "ATAN2"(Y:=#X.im,X:=#X.re);

   #CLOG := #temp_complex;

   (* revision history
   hm  21. feb 2008    rev 1.0
       original version

   hm  20. apr. 2008   rev 1.1
       use ATAN2 instead of ATAN
   *)
END_FUNCTION

FUNCTION "CMUL" : "COMPLEX"   // FC133, SCL
TITLE = CMUL
{ S7_Optimized_Access := 'FALSE' }
AUTHOR : hugo
FAMILY : CMATH
NAME : CMUL
VERSION : 1.0
// this function multiplies two complex numbers
// 
// uses: COMPLEX [UDT2]
   VAR_INPUT
      X : "COMPLEX";
      Y : "COMPLEX";
   END_VAR
   VAR_TEMP
      temp_CMUL : "COMPLEX";
   END_VAR
BEGIN


     #temp_CMUL.re := #X.re * #Y.re - #X.im * #Y.im;
     #temp_CMUL.im := #X.re * #Y.im + #X.im * #Y.re;

     #CMUL := #temp_CMUL;

   (* revision history
   hm  21. feb 2008  rev 1.0
     original version

   *)
END_FUNCTION

FUNCTION "CPOL" : "COMPLEX"   // FC134, SCL
TITLE = CPOL
{ S7_Optimized_Access := 'FALSE' }
AUTHOR : hugo
FAMILY : CMATH
NAME : CPOL
VERSION : 1.0
// this function creates a complex numbers for the polar form with the inputs L (length) an A for Angle.
// 
// uses: COMPLEX [UDT2]
   VAR_INPUT
      L : Real;
      "A" : Real;
   END_VAR
   VAR_TEMP
      temp_CPOL : "COMPLEX";
   END_VAR
BEGIN


     #temp_CPOL.re := #L * COS(#"A");
     #temp_CPOL.im := #L * SIN(#"A");

     #CPOL := #temp_CPOL;

   (* revision history
   hm  21. feb 2008  rev 1.0
     original version

   *)
END_FUNCTION

FUNCTION "CPOW" : "COMPLEX"   // FC135, SCL
TITLE = CPOW
{ S7_Optimized_Access := 'FALSE' }
AUTHOR : hugo
FAMILY : CMATH
NAME : CPOW
VERSION : 1.0
// this function calculates the complex power function x to the power of y
// 
// uses: COMPLEX [UDT2]
//       CEXP [FC130]
//       CMUL [FC133]
//       CLOG [FC132]
//       HYPOT [FC89] 
//       ATAN2 [FC58]
   VAR_INPUT
      X : "COMPLEX";
      Y : "COMPLEX";
   END_VAR
   VAR_TEMP
      temp_X : "COMPLEX";
      temp_Y : "COMPLEX";
      temp_CPOW : "COMPLEX";
   END_VAR
BEGIN


     #temp_X := #X;
     #temp_Y := #Y;

     #temp_CPOW := "CEXP"("CMUL"(Y:=#temp_Y,X:="CLOG"(#temp_X)));

     #CPOW := #temp_CPOW;

   (* revision history
   hm  21. feb 2008  rev 1.0
     original version

   *)
END_FUNCTION

FUNCTION "CSET" : "COMPLEX"   // FC136, SCL
TITLE = CSET
{ S7_Optimized_Access := 'FALSE' }
AUTHOR : hugo
FAMILY : CMATH
NAME : CSET
VERSION : 1.0
// this function creates a complex number from two real inputs
// 
// uses: COMPLEX [UDT2]
   VAR_INPUT
      RE : Real;
      IM : Real;
   END_VAR
   VAR_TEMP
      temp_CSET : "COMPLEX";
   END_VAR
BEGIN


     #temp_CSET.re := #RE;
     #temp_CSET.im := #IM;

     #CSET := #temp_CSET;

   (* revision history
   hm  21. feb 2008  rev 1.0
     original version

   *)
END_FUNCTION

FUNCTION "CSIN" : "COMPLEX"   // FC137, SCL
TITLE = CSIN
{ S7_Optimized_Access := 'FALSE' }
AUTHOR : hugo
FAMILY : CMATH
NAME : CSIN
VERSION : 1.0
// this function calculates the sinus function of a complex number
// 
// uses: COMPLEX [UDT2]
//       COSH [FC69]
//       SINH [FC111]
   VAR_INPUT
      X : "COMPLEX";
   END_VAR
   VAR_TEMP
      temp_CSIN : "COMPLEX";
   END_VAR
BEGIN


     #temp_CSIN.re := "COSH"(#X.im) * SIN(#X.re);
     #temp_CSIN.im := "SINH"(#X.im) * COS(#X.re);

     #CSIN := #temp_CSIN;

   (* revision history
   hm  21. feb 2008  rev 1.0
     original version

   *)
END_FUNCTION

FUNCTION "CSINH" : "COMPLEX"   // FC138, SCL
TITLE = CSINH
{ S7_Optimized_Access := 'FALSE' }
AUTHOR : hugo
FAMILY : CMATH
NAME : CSINH
VERSION : 1.0
// this function calculates the sinus function of a complex number
//  
// uses: COMPLEX [UDT2]
//       SINH [FC111]
//       COSH [FC69]
   VAR_INPUT
      X : "COMPLEX";
   END_VAR
   VAR_TEMP
      temp_CSINH : "COMPLEX";
   END_VAR
BEGIN


     #temp_CSINH.re := "SINH"(#X.re) * COS(#X.im);
     #temp_CSINH.im := "COSH"(#X.re) * SIN(#X.im);

     #CSINH := #temp_CSINH;

   (* revision history
   hm  21. feb 2008  rev 1.0
     original version

   *)
END_FUNCTION

FUNCTION "CSQRT" : "COMPLEX"   // FC139, SCL
TITLE = CSQRT
{ S7_Optimized_Access := 'FALSE' }
AUTHOR : hugo
FAMILY : CMATH
NAME : CSQRT
VERSION : 1.0
// this function calculates the complex sqare root
// 
// uses: COMPLEX [UDT2]
//       HYPOT [FC89]
//       SGN [FC106]
   VAR_INPUT
      X : "COMPLEX";
   END_VAR
   VAR_TEMP
      temp : Real;
      temp_complex : "COMPLEX";
   END_VAR
BEGIN


     #temp := "HYPOT"(X:=#X.re,Y:=#X.im);
     #temp_complex.re :=  SQRT(0.5 * (#temp + #X.re));
     #temp_complex.im :=  "SGN"(#X.im) * SQRT(0.5 * (#temp - #X.re));

     #CSQRT := #temp_complex;

   (* revision history
   hm  21. feb 2008  rev 1.0
     original version

   *)
END_FUNCTION

FUNCTION "CSUB" : "COMPLEX"   // FC140, SCL
TITLE = CSUB
{ S7_Optimized_Access := 'FALSE' }
AUTHOR : hugo
FAMILY : CMATH
NAME : CSUB
VERSION : 1.0
// this function subtracts two complex numbers
// 
// uses: COMPLEX [UDT2]
   VAR_INPUT
      X : "COMPLEX";
      Y : "COMPLEX";
   END_VAR
   VAR_TEMP
      temp_CSUB : "COMPLEX";
   END_VAR
BEGIN


     #temp_CSUB.re := #X.re - #Y.re;
     #temp_CSUB.im := #X.im - #Y.im;

     #CSUB := #temp_CSUB;

   (* revision history
   hm  21. feb 2008  rev 1.0
     original version

   *)
END_FUNCTION

FUNCTION "CTAN" : "COMPLEX"   // FC141, SCL
TITLE = CTAN
{ S7_Optimized_Access := 'FALSE' }
AUTHOR : hugo
FAMILY : CMATH
NAME : CTAN
VERSION : 1.1
// this function calculates the tangens function of a complex number
//  
// uses: COMPLEX [UDT2]
//       COSH [FC69]
//       SINH [FC111]
   VAR_INPUT
      X : "COMPLEX";
   END_VAR
   VAR_TEMP
      temp : Real;
      xi2 : Real;
      xr2 : Real;
      tCTAN : "COMPLEX";
   END_VAR
BEGIN


   #xi2 := 2.0 * #X.im;
   #xr2 := 2.0 * #X.re;
   #temp := 1.0 / (COS(#xr2) + "COSH"( #xi2));
   #tCTAN.re := #temp * SIN(#xr2);
   #tCTAN.im := #temp * "SINH"(#xi2);

   #CTAN := #tCTAN;


   (* revision history
   hm  21. feb 2008    rev 1.0
       original version

   hm  10. mar 2009    rev 1.1
       faster code
   *)
END_FUNCTION

FUNCTION "CTANH" : "COMPLEX"   // FC142, SCL
TITLE = CTANH
{ S7_Optimized_Access := 'FALSE' }
AUTHOR : hugo
FAMILY : CMATH
NAME : CTANH
VERSION : 1.1
// this function calculates the complex hyperbolictangens
// 
// uses: COMPLEX [UDT2]
//       COSH [FC69]
//       SINH [FC111]
   VAR_INPUT
      X : "COMPLEX";
   END_VAR
   VAR_TEMP
      temp : Real;
      xi2 : Real;
      xr2 : Real;
      tCTANH : "COMPLEX";
   END_VAR
BEGIN


   #xi2 := 2.0 * #X.im;
   #xr2 := 2.0 * #X.re;
   #temp := 1.0 / ("COSH"(#xr2) + COS(#xi2));
   #tCTANH.re := #temp * "SINH"(#xr2);
   #tCTANH.im := #temp * SIN(#xi2);

   #CTANH := #tCTANH;


   (* revision history
   hm  21. feb 2008    rev 1.0
       original version

   hm  10. mar. 2009   rev 1.1 
       new faster code

   *)
END_FUNCTION

// ===== PLC "Mathematical Geometry"  Unspecific CPU S7 300 =====

VAR_GLOBAL CONSTANT   // PLC tag table "STEP7 classic symbols"
   "PI2" : Real := 6.283185307179586476;   // PI * 2
   "PI" : Real := 3.14159265358979323846264338327950288;   // Kreiszahl PI
END_VAR

FUNCTION "FLOOR2" : DInt   // FC82, SCL
TITLE = FLOOR2
{ S7_Optimized_Access := 'FALSE' }
AUTHOR : hugo
FAMILY : MATH
NAME : FLOOR2
VERSION : 1.1
// This is a rounding function which returns the biggest possible integer which is less or equal to X.
// floor2(3.14) = 3
// floor2(-3.14) = -4
   VAR_INPUT
      X : Real;
   END_VAR
BEGIN


   #FLOOR2 := REAL_TO_DINT(#X);
   IF DINT_TO_REAL(#FLOOR2) > #X THEN
     #FLOOR2 := #FLOOR2 - 1;
   END_IF;

   (* revision history
   hm  21. mar. 2008   rev 1.0
       originlal version

   hm  4. apr. 2008    rev 1.1
       added type conversion to avoid warnings under codesys 3.0
   *)
END_FUNCTION

FUNCTION "MODR" : Real   // FC97, SCL
TITLE = MODR
{ S7_Optimized_Access := 'FALSE' }
AUTHOR : hugo
FAMILY : MATH
NAME : MODR
VERSION : 1.5
// this is a modulo funtion for real numbers
// modr(5.5,2.5) = 0.5
// 
// uses: FLOOR2 [FC82]
   VAR_INPUT
      IN : Real;
      DIVI : Real;
   END_VAR
BEGIN


   IF #DIVI = 0.0 THEN
       #MODR := 0.0;
   ELSE
       #MODR := #IN - DINT_TO_REAL("FLOOR2"(#IN / #DIVI)) * #DIVI;
   END_IF;


   (* revision history

   hm  4. aug.2006     rev 1.0

   hm  28. jan.2007   rev 1.1
       modr(x,0) will deliver the result 0

   hm  21. mar 2008    rev 1.2
       use D_trunc for compatibility reasons

   hm  4. apr. 2008    rev 1.3
       added type conversion to avoid warnings under codesys 3.0

   hm  31. oct. 2008   rev 1.4
       changed algorithm to the more common version using floor instead of TRUNC

   hm  10. mar. 2009   rev 1.5
       real constants updated to new systax using dot

   *)
END_FUNCTION

FUNCTION "RAD" : Real   // FC100, SCL
TITLE = RAD
{ S7_Optimized_Access := 'FALSE' }
AUTHOR : hugo
FAMILY : MATH
NAME : RAD
VERSION : 1.2
// this function converts Radiant to degrees
// 
// uses: MODR [FC97]
//       FLOOR2 [FC82]
   VAR_INPUT
      deg : Real;
   END_VAR
BEGIN


   #RAD := "MODR"(IN:=0.0174532925199433 * #deg,DIVI:="PI2");

   (*  Enfällt da der Zugriff auf Datenbaustein länger dauert
       RAD := MODR(0.0174532925199433 * DEG, math.PI2);
   *)

   (* revision history
   hm  4. aug 2006     rev 1.0
       original version

   hm  16. oct 2007    rev 1.1
       added modr statement which prohibits rad to become bigger than 2PI

   hm  18. oct 2008    rev 1.2
       using math constants

   *)
END_FUNCTION

FUNCTION "CIRCLE_A" : Real   // FC155, SCL
TITLE = CIRCLE_A
{ S7_Optimized_Access := 'FALSE' }
AUTHOR : hugo
FAMILY : GEOMETRY
NAME : CIRCLE_A
VERSION : 1.2
// circle_A calculates the Area of a circle segement if ax = 360 the whole circle is calculated
   VAR_INPUT
      rx : Real;
      ax : Real;
   END_VAR
BEGIN


     #CIRCLE_A := #rx * #rx * 8.726646E-3 * #ax;

   (* revision histroy
   hm  16. oct 2007  rev 1.0
     original version

   hm  4. dec 2007   rev 1.1
     changed code for better performance

   hm  22. feb 2008  rev 1.2
     improved performance
   *)
END_FUNCTION

FUNCTION "CIRCLE_C" : Real   // FC156, SCL
TITLE = CIRCLE_C
{ S7_Optimized_Access := 'FALSE' }
AUTHOR : hugo
FAMILY : GEOMETRY
NAME : CIRCLE_C
VERSION : 1.1
// circle_C calculates the Circumference of a circle  if ax = 360 the whole circle is calculated
   VAR_INPUT
      Rx : Real;
      Ax : Real;
   END_VAR
BEGIN


     #CIRCLE_C := 1.7453293E-2 * #Rx * #Ax;

   (* revision histroy
   hm  16. oct 2007  rev 1.0
     original version

   hm  22. feb 2008  rev 1.1
     improved performance
   *)
END_FUNCTION

FUNCTION "CONE_V" : Real   // FC157, SCL
TITLE = CONE_V
{ S7_Optimized_Access := 'FALSE' }
AUTHOR : hugo
FAMILY : GEOMETRY
NAME : CONE_V
VERSION : 1.2
// cone_V calculates the Volume of a cone
   VAR_INPUT
      rx : Real;
      hx : Real;
   END_VAR
BEGIN


     #CONE_V := 1.047197551 * #rx * #rx * #hx;

   (* revision histroy
   hm  17. oct 2007  rev 1.0
     original version

   hm  4. dec 2007   rev 1.1
     changed code for better performance

   hm  22. feb 2008  rev 1.2
     changed code for better performance
   *)
END_FUNCTION

FUNCTION "ELLIPSE_A" : Real   // FC158, SCL
TITLE = ELLIPSE_A
{ S7_Optimized_Access := 'FALSE' }
AUTHOR : hugo
FAMILY : GEOMETRY
NAME : ELLIPS_A
VERSION : 1.1
// ellipse_A calculates the Area of an ellipe based on the two radians R1 and R2
   VAR_INPUT
      R1 : Real;
      R2 : Real;
   END_VAR
BEGIN


   #ELLIPSE_A := "PI" * #R1 * #R2;

   (*  Käse!
       ELLIPSE_A := math.PI * R1 * R2;
   *)

   (* revision histroy
   hm  16. oct 2007    rev 1.0
       original version

   hm  18. oct. 2008   rev 1.1
       using math constants
   *)
END_FUNCTION

FUNCTION "ELLIPSE_C" : Real   // FC159, SCL
TITLE = ELLIPSE_C
{ S7_Optimized_Access := 'FALSE' }
AUTHOR : hugo
FAMILY : GEOMETRY
NAME : ELLIPS_C